// TIA Portal project "FS-DS-09" (V16)
// C100锁螺丝机

(* hardware
DEVICE "S7-1200 station_1"  S7-1200 Station
   slot 0: "Rack_0"  S7-1200 Rack  Rack  V1.0
   slot 1: "FS-DS-09"  CPU 1214C DC/DC/DC  6ES7 214-1AG40-0XB0  V4.4
   slot 2: "DI 16/DQ 16x24VDC_1"  6ES7 223-1BL32-0XB0  V2.0
   slot 3: "DI 8/DQ 8x24VDC_1"  6ES7 223-1BH32-0XB0  V2.0
DEVICE "HMI_1"  KTP700 Basic PN
   slot 0: "HMI_1"  KTP700 Basic PN  6AV2 123-2GB03-0AX0  16.0.0.0
   slot 1: "HMI_RT_1"  KTP700 Basic PN  6AV2 123-2GB03-0AX0  16.0.0.0
   slot 5: "HMI_1.IE_CP_1"  PROFINET Interface  16.0.0.0
      slot 1: "PROFINET Interface_1"  PROFINET Interface
         slot 1: "Port_1"  Port
DEVICE "GSD device_1"  GSD.Device.PN
   slot 0: "机架"  Rack  V1.0
   slot 0: "hj6300"  HJ6300-PN-hj6302-2789  HJ6300-PN  -V1.2
      slot 0: "HJ6300-PN-hj6302-2789"  HJ6300-PN-hj6302-2789
      slot 1: "Interface"  Interface
         slot 1: "Port1"  Port1
         slot 2: "Port2"  Port2
      slot 1: "X逻辑输入 COM1/addr=2/reg=17410_1"  X逻辑输入 COM1/addr=2/reg=17410
         slot 0: "X逻辑输入 COM1/addr=2/reg=17410"  X逻辑输入 COM1/addr=2/reg=17410
      slot 2: "Y逻辑输入 COM1/addr=3/reg=17410_1"  Y逻辑输入 COM1/addr=3/reg=17410
         slot 0: "Y逻辑输入 COM1/addr=3/reg=17410"  Y逻辑输入 COM1/addr=3/reg=17410
      slot 3: "Z逻辑输入 COM1/addr=4/reg=17410_1"  Z逻辑输入 COM1/addr=4/reg=17410
         slot 0: "Z逻辑输入 COM1/addr=4/reg=17410"  Z逻辑输入 COM1/addr=4/reg=17410
      slot 4: "x读取错误编号 COM1/addr=2/reg=24577_1"  x读取错误编号 COM1/addr=2/reg=24577
         slot 0: "x读取错误编号 COM1/addr=2/reg=24577"  x读取错误编号 COM1/addr=2/reg=24577
      slot 5: "y读取错误编号 COM1/addr=3/reg=24577_1"  y读取错误编号 COM1/addr=3/reg=24577
         slot 0: "y读取错误编号 COM1/addr=3/reg=24577"  y读取错误编号 COM1/addr=3/reg=24577
      slot 6: "z读取错误编号 COM1/addr=4/reg=24577_1"  z读取错误编号 COM1/addr=4/reg=24577
         slot 0: "z读取错误编号 COM1/addr=4/reg=24577"  z读取错误编号 COM1/addr=4/reg=24577
      slot 7: "x读取速度 COM1/addr=2/reg=19718_1"  x读取速度 COM1/addr=2/reg=19718
         slot 0: "x读取速度 COM1/addr=2/reg=19718"  x读取速度 COM1/addr=2/reg=19718
      slot 8: "y读取速度 COM1/addr=3/reg=19718_1"  y读取速度 COM1/addr=3/reg=19718
         slot 0: "y读取速度 COM1/addr=3/reg=19718"  y读取速度 COM1/addr=3/reg=19718
      slot 9: "z读取速度 COM1/addr=4/reg=19718_1"  z读取速度 COM1/addr=4/reg=19718
         slot 0: "z读取速度 COM1/addr=4/reg=19718"  z读取速度 COM1/addr=4/reg=19718
      slot 10: "x轴逻辑输出 COM1/addr=2/reg=17481_1"  x轴逻辑输出 COM1/addr=2/reg=17481
         slot 0: "x轴逻辑输出 COM1/addr=2/reg=17481"  x轴逻辑输出 COM1/addr=2/reg=17481
      slot 11: "y轴逻辑输出 COM1/addr=3/reg=17481_1"  y轴逻辑输出 COM1/addr=3/reg=17481
         slot 0: "y轴逻辑输出 COM1/addr=3/reg=17481"  y轴逻辑输出 COM1/addr=3/reg=17481
      slot 12: "z轴逻辑输出 COM1/addr=4/reg=17481_1"  z轴逻辑输出 COM1/addr=4/reg=17481
         slot 0: "z轴逻辑输出 COM1/addr=4/reg=17481"  z轴逻辑输出 COM1/addr=4/reg=17481
      slot 14: "Alarm Data Module_1"  Alarm Data Module
         slot 0: "Alarm Data SubModule"  Alarm Data SubModule
*)

// ===== PLC "FS-DS-09"  CPU 1214C DC/DC/DC =====

VAR_GLOBAL   // PLC tag table "默认变量表"
   "Clock_Byte" AT %MB0 : Byte;
   "Clock_10Hz" AT %M0.0 : Bool;
   "Clock_5Hz" AT %M0.1 : Bool;
   "Clock_2.5Hz" AT %M0.2 : Bool;
   "Clock_2Hz" AT %M0.3 : Bool;
   "Clock_1.25Hz" AT %M0.4 : Bool;
   "Clock_1Hz" AT %M0.5 : Bool;
   "Clock_0.625Hz" AT %M0.6 : Bool;
   "Clock_0.5Hz" AT %M0.7 : Bool;
   "System_Byte" AT %MB1 : Byte;
   "FirstScan" AT %M1.0 : Bool;
   "DiagStatusUpdate" AT %M1.1 : Bool;
   "AlwaysTRUE" AT %M1.2 : Bool;
   "AlwaysFALSE" AT %M1.3 : Bool;
   "Tag_1" AT %M4.0 : Bool;
   "Tag_2" AT %M6.0 : Bool;
   "Tag_3" AT %M5.0 : Bool;
   "Tag_4" AT %M200.0 : Bool;
   "Tag_5" AT %M200.1 : Bool;
   "Tag_6" AT %M30.0 : Bool;
   "Tag_7" AT %M30.1 : Bool;
   "Tag_8" AT %M60.0 : Bool;
   "Tag_9" AT %M20.0 : Bool;
   "Tag_10" AT %M50.0 : Bool;
   "Tag_11" AT %M50.1 : Bool;
   "Tag_12" AT %M50.2 : Bool;
END_VAR

VAR_GLOBAL   // PLC tag table "输入"
   "操作面板急停" AT %I0.0 : Bool;
   "回原位" AT %I0.1 : Bool;
   "启动按钮" AT %I0.2 : Bool;
   "停止按钮" AT %I0.3 : Bool;
   "手动/自动" AT %I0.4 : Bool;
   "按钮盒急停" AT %I0.5 : Bool;
   "左启动" AT %I0.6 : Bool;
   "右启动" AT %I0.7 : Bool;
   "备用" AT %I1.0 : Bool;
   "光幕" AT %I1.1 : Bool;
   "Y1供料器有料" AT %I1.2 : Bool;
   "Y2供料器有料" AT %I1.3 : Bool;
   "1#工装产品信号" AT %I1.4 : Bool;
   "2#工装产品信号" AT %I1.5 : Bool;
   "气夹气缸到位2" AT %I2.0 : Bool;
   "气夹气缸到位1" AT %I2.1 : Bool;
   "工具错误" AT %I2.2 : Bool;
   "工具拧紧OK" AT %I2.3 : Bool;
   "工具拧紧NG" AT %I2.4 : Bool;
   "工具准备好" AT %I2.5 : Bool;
   "工具运行" AT %I2.6 : Bool;
   "气源压力检测" AT %I2.7 : Bool;
   "光栅屏蔽对射开关" AT %I3.0 : Bool;
   "吸附信号" AT %I3.1 : Bool;
   "电批下压气缸下压信号" AT %I3.2 : Bool;
   "安全门" AT %I3.3 : Bool;
   "回原位中" AT %I3.4 : Bool;
   "回原位完成" AT %I3.5 : Bool;
   "X轴故障报警" AT %I3.6 : Bool;
   "Y轴故障报警" AT %I3.7 : Bool;
   "Z轴故障报警" AT %I4.0 : Bool;
   "运动控制卡完成/释放夹紧气缸" AT %I4.1 : Bool;
   "备用_3" AT %I4.2 : Bool;
   "备用_4" AT %I4.3 : Bool;
   "备用_5" AT %I4.4 : Bool;
   "备用_6" AT %I4.5 : Bool;
   "备用_7" AT %I4.6 : Bool;
   "备用_8" AT %I4.7 : Bool;
END_VAR

VAR_GLOBAL   // PLC tag table "输出"
   "三色灯黄色" AT %Q0.0 : Bool;
   "三色灯绿色" AT %Q0.1 : Bool;
   "三色灯红色" AT %Q0.2 : Bool;
   "三色灯蜂鸣器" AT %Q0.3 : Bool;
   "绿色半球指示灯" AT %Q0.4 : Bool;
   "红色半球指示灯" AT %Q0.5 : Bool;
   "运动控制卡任务选择1" AT %Q0.6 : Bool;
   "运动控制卡任务选择2" AT %Q0.7 : Bool;
   "运动控制卡任务选择3" AT %Q1.0 : Bool;
   "运动控制卡任务选择4" AT %Q1.1 : Bool;
   "运动控制卡任务选择5" AT %Q2.0 : Bool;
   "Y1供料器有料输出" AT %Q2.1 : Bool;
   "Y2供料器有料输出" AT %Q2.2 : Bool;
   "运动控制卡启动" AT %Q2.3 : Bool;
   "运动控制卡复位" AT %Q2.4 : Bool;
   "运动控制卡紧急停止" AT %Q2.5 : Bool;
   "运动控制卡停止" AT %Q2.6 : Bool;
   "吸取螺丝电磁阀" AT %Q2.7 : Bool;
   "下压气缸电磁阀" AT %Q3.0 : Bool;
   "工装电磁铁" AT %Q3.1 : Bool;
   "光栅报警" AT %Q3.2 : Bool;
   "伺服复位" AT %Q3.3 : Bool;
   "电批急停" AT %Q3.4 : Bool;
   "电批测试启动" AT %Q3.5 : Bool;
   "FFU" AT %Q3.6 : Bool;
   "照明" AT %Q3.7 : Bool;
   "左启动指示灯" AT %Q4.0 : Bool;
   "右启动指示灯" AT %Q4.1 : Bool;
   "夹紧气缸夹紧" AT %Q4.2 : Bool;
   "伺服报警" AT %Q4.3 : Bool;
   "备用_5(1)" AT %Q4.4 : Bool;
   "备用_6(1)" AT %Q4.5 : Bool;
   "备用_7(1)" AT %Q4.6 : Bool;
   "备用_8(1)" AT %Q4.7 : Bool;
END_VAR

VAR_GLOBAL   // PLC tag table "伺服变量"
   "负方向x" AT %I6.2 : Bool;
   "正方向x" AT %I6.3 : Bool;
   "准备OKx" AT %I42.0 : Bool;
   "故障报警x" AT %I42.1 : Bool;
   "故障代码x" AT %ID17 : DWord;
   "负方向y" AT %I10.2 : Bool;
   "正方向y" AT %I10.3 : Bool;
   "准备OKy" AT %I46.0 : Bool;
   "故障报警y" AT %I46.1 : Bool;
   "故障代码y" AT %ID21 : DWord;
   "负方向z" AT %I14.2 : Bool;
   "正方向z" AT %I14.3 : Bool;
   "准备OKz" AT %I50.0 : Bool;
   "故障报警z" AT %I50.1 : Bool;
   "故障代码z" AT %ID25 : DWord;
END_VAR

TYPE "hengkong"
   STRUCT
      DATA : Struct
         X轴原位 : Bool;
         Y轴原位 : Bool;
         Z轴原位 : Bool;
         Y1供料器有料 : Bool;
         Y2供料器有料 : Bool;
         备用 : Bool;
         任务选择1 : Bool;
         任务选择2 : Bool;
         启动 : Bool;
         回原位 : Bool;
         急停 : Bool;
         OK : Bool;
         光幕和门控报警 : Bool;
         任务选择3 : Bool;
         任务选择4 : Bool;
         任务选择5 : Bool;
         负压传感器 : Bool;
         备用_1 : Bool;
         备用_2 : Bool;
         备用_3 : Bool;
         备用_4 : Bool;
         下压气缸原位 : Bool;
         备用_5 : Bool;
         停止 : Bool;
         吸取螺丝信号 : Bool;
         回原位成功 : Bool;
         回原位中 : Bool;
         下压气缸信号 : Bool;
         备用_6 : Bool;
         认螺帽反转 : Bool;
         备用_7 : Bool;
         备用_8 : Bool;
         任务选择0 : Bool;
         任务选择6 : Bool;
         任务选择7 : Bool;
         备用_9 : Bool;
         启动电批 : Bool;
         备用_10 : Bool;
         备用_11 : Bool;
         备用_12 : Bool;
         获取X轴当前坐标 : LReal;
         获取Y轴当前坐标 : LReal;
         获取Z轴当前坐标 : LReal;
         获取Y2轴当前坐标 : LReal;
         完成螺丝数量 : LReal;
         完成产品数量 : LReal;
         产品合格率 : Word;
         螺丝孔加工完成情况查询 : Word;
         设备报警状态查询 : Word;
         左机加工完成情况查询 : Word;
         右机加工完成情况查询 : Word;
         允许运行指令 : Word;
         从机地址 : Word;
         智能电批任务号 : Word;
         电批加工NG时处理指令 : Word;
      END_STRUCT;
   END_STRUCT;
END_TYPE

TYPE "UDPP"
   STRUCT
      加工文件名称 : String;
      加工文件编号 : Int;
      加工螺丝数量 : Int;
   END_STRUCT;
END_TYPE

TYPE "产品"
   STRUCT
      配方 : Struct
         示教器程序号 : Int;
         产品名称 : String;
      END_STRUCT;
   END_STRUCT;
END_TYPE

DATA_BLOCK "count_DB"   // DB18
{ S7_Optimized_Access := 'TRUE' }
VERSION : 0.1
// stored: InstanceOfName count
"count"
BEGIN
END_DATA_BLOCK

// folder: Alarm

DATA_BLOCK "Alarm FB_DB"   // DB5
{ S7_Optimized_Access := 'TRUE' }
VERSION : 0.1
// stored: InstanceOfName Alarm FB
"Alarm FB"
BEGIN
END_DATA_BLOCK

// folder: Control

DATA_BLOCK "Control_DB"   // DB6
{ S7_Optimized_Access := 'TRUE' }
VERSION : 0.1
// stored: InstanceOfName Control FB
"Control FB"
BEGIN
END_DATA_BLOCK

DATA_BLOCK "Start_DB"   // DB9
{ S7_Optimized_Access := 'TRUE' }
VERSION : 0.1
// stored: InstanceOfName Start
"Start"
BEGIN
END_DATA_BLOCK

DATA_BLOCK "吐钉模式"   // DB20
{ S7_Optimized_Access := 'TRUE' }
VERSION : 0.1
   VAR
      吐钉模式 : Bool;
      下压气缸复位信号 : Bool;
      启动就绪 : Bool;
   END_VAR
BEGIN
END_DATA_BLOCK

// folder: DATA

DATA_BLOCK "IO"   // DB1
{ S7_Optimized_Access := 'FALSE' }
VERSION : 0.1
   VAR
      IN : Array[0..40] of Bool;
      OUT : Array[0..40] of Bool;
   END_VAR
BEGIN
   // IN[0] : 操作面板急停
   // IN[1] : 回原位
   // IN[2] : 启动按钮
   // IN[3] : 停止按钮
   // IN[4] : 手动/自动
   // IN[5] : 按钮盒急停
   // IN[6] : 左启动
   // IN[7] : 右启动
   // IN[8] : 备用
   // IN[9] : 光幕
   // IN[10] : Y1供料器有料
   // IN[11] : Y2供料器有料
   // IN[12] : 1#工装产品信号
   // IN[13] : 2#工装产品信号
   // IN[14] : 气夹气缸到位2
   // IN[15] : 气夹气缸到位1
   // IN[16] : 工具错误
   // IN[17] : 工具拧紧OK
   // IN[18] : 工具拧紧NG
   // IN[19] : 工具准备好
   // IN[20] : 工具运行
   // IN[21] : 气源压力检测
   // IN[22] : 光栅屏蔽对射开关
   // IN[23] : 吸附信号
   // IN[24] : 电批下压气缸下压信号
   // IN[25] : 安全门
   // IN[26] : 回原位中
   // IN[27] : 回原位完成
   // IN[28] : X轴故障报警
   // IN[29] : Y轴故障报警
   // IN[30] : Z轴故障报警
   // IN[31] : 运动控制卡完成/释放夹紧气缸
   // IN[32] : 备用_3
   // IN[33] : 备用_4
   // IN[34] : 备用_5
   // IN[35] : 备用_6
   // IN[36] : 备用_7
   // IN[37] : 备用_8
   // OUT[0] : 三色灯黄色
   // OUT[1] : 三色灯绿色
   // OUT[2] : 三色灯红色
   // OUT[3] : 三色灯蜂鸣器
   // OUT[4] : 绿色半球指示灯
   // OUT[5] : 红色半球指示灯
   // OUT[6] : 运动控制卡任务选择1
   // OUT[7] : 运动控制卡任务选择2
   // OUT[8] : 运动控制卡任务选择3
   // OUT[9] : 运动控制卡任务选择4
   // OUT[10] : 运动控制卡任务选择5
   // OUT[11] : Y1供料器有料输出
   // OUT[12] : Y2供料器有料输出
   // OUT[13] : 运动控制卡启动
   // OUT[14] : 运动控制卡复位
   // OUT[15] : 运动控制卡紧急停止
   // OUT[16] : 运动控制卡停止
   // OUT[17] : 吸取螺丝电磁阀
   // OUT[18] : 下压气缸电磁阀
   // OUT[19] : 工装电磁铁
   // OUT[20] : 光栅报警
   // OUT[21] : 伺服复位
   // OUT[22] : 电批急停
   // OUT[23] : 电批测试启动
   // OUT[24] : FFU
   // OUT[25] : 照明
   // OUT[26] : 左启动指示灯
   // OUT[27] : 右启动指示灯
   // OUT[28] : 夹紧气缸夹紧
   // OUT[29] : 伺服报警
   // OUT[30] : 备用_5(1)
   // OUT[31] : 备用_6(1)
   // OUT[32] : 备用_7(1)
   // OUT[33] : 备用_8(1)
END_DATA_BLOCK

DATA_BLOCK "HengKongMC"   // DB2
{ S7_Optimized_Access := 'FALSE' }
VERSION : 0.1
   VAR
      输入 : Struct   // R/W 01/05/0F
         X轴原位 : Bool;   // 4096
         Y轴原位 : Bool;   // 4097
         Z轴原位 : Bool;   // 4098
         X4备用 : Bool;   // 4099
         Y2供料器有料 : Bool;   // 4100
         电批启动 : Bool;   // 4101
         任务选择1 : Bool;   // 4102
         任务选择2 : Bool;   // 4103
         启动 : Bool;   // 4104
         回原位 : Bool;   // 4105
         急停 : Bool;   // 4106
         OK : Bool;   // 4107
         光幕和门控报警 : Bool;   // 4108
         任务选择3 : Bool;   // 4109
         任务选择4 : Bool;   // 4110
         任务选择5 : Bool;   // 4111
         负压传感器 : Bool;   // 4112
         Y1供料器有料 : Bool;   // 4113
         X19 : Bool;   // 4114
         X20 : Bool;   // 4115
         X21 : Bool;   // 4116
         下压气缸原位 : Bool;   // 4117
         X23 : Bool;   // 4118
         停止 : Bool;   // 4119
      END_STRUCT;
      输出 : Struct   // R/W 01/05/0F
         吸取螺丝信号 : Bool;   // 4176
         回原位成功 : Bool;   // 4177
         回原位中 : Bool;   // 4178
         下压气缸信号 : Bool;   // 4179
         Y5 : Bool;   // 4180
         认螺帽反转 : Bool;   // 4181
         运动控制卡完成信号 : Bool;   // 4182
         Y8 : Bool;   // 4183
         任务选择0 : Bool;   // 4184
         任务选择1 : Bool;   // 4185
         任务选择2 : Bool;   // 4186
         Y12 : Bool;   // 4187
         启动电批 : Bool;   // 4188
         Y14 : Bool;   // 4189
         回原位标志位 : Bool;   // 4190
         Y16 : Bool;   // 4191
      END_STRUCT;
      hengkong : Struct   // 运动控制板卡
         获取X轴当前坐标 : LReal;
         获取Y轴当前坐标 : LReal;
         获取Z轴当前坐标 : LReal;
         获取Y2轴当前坐标 : LReal;
         完成螺丝数量 : Int;
         完成产品数量 : Int;
         产品合格率 : Int;
         螺丝孔加工完成情况查询 : Word;
         设备报警状态查询 : Word;
         左机加工完成情况查询 : Word;
         右机加工完成情况查询 : Word;
         报警异常号 : Int;
         光标处运行标志 : Int;
         当前程序所在行号 : Int;
      END_STRUCT;
   END_VAR
BEGIN
END_DATA_BLOCK

DATA_BLOCK "Alarm"   // DB4
{ S7_Optimized_Access := 'FALSE' }
VERSION : 0.1
   VAR
      运动控制板卡螺丝加工完成情况昂查询 : String;
      运动控制板卡设备报警状态查询 : String;
      运动控制板卡报警 : Bool;
      设备气源压力低报警 : Bool;
      面板急停报警 : Bool;
      操作面板急停报警 : Bool;
      安全门报警 : Bool;
      光幕报警 : Bool;
      回原位超时报警 : Bool;
      Y1供料器超时报警 : Bool;
      Y2供料器超时报警 : Bool;
      工装产品检测1无件报警 : Bool;
      工装产品检测2无件报警 : Bool;
      气缸夹紧1夹紧超时 : Bool;
      气缸夹紧2夹紧超时 : Bool;
      丹尼克尔错误报警 : Bool;
      一级报警 : Bool;
      二级报警 : Bool;
      下压气缸故障 : Bool;
      打螺丝延时过小 : Bool;
      真空检测失败 : Bool;
      吸取螺丝失败 : Bool;
      分料超时 : Bool;
      夹紧气缸故障FB运行前未复位 : Bool;
      下压气缸不在原位 : Bool;
      X轴故障报警 : Bool;
      Y轴故障报警 : Bool;
      Z轴故障报警 : Bool;
   END_VAR
BEGIN
END_DATA_BLOCK

DATA_BLOCK "Blocking function"   // DB7
{ S7_Optimized_Access := 'FALSE' }
VERSION : 0.1
   VAR
      Y1供料器报警屏蔽 : Bool;
      Y2供料器报警屏蔽 : Bool;
      工装产品检测1屏蔽 : Bool;
      工装产品检测2屏蔽 : Bool;
      夹紧气缸1夹紧屏蔽 : Bool;
      夹紧气缸2夹紧屏蔽 : Bool;
      上位机屏蔽 : Bool;
      安全门屏蔽 : Bool;
      光幕屏蔽 : Bool;
   END_VAR
BEGIN
END_DATA_BLOCK

DATA_BLOCK "Control"   // DB8
{ S7_Optimized_Access := 'FALSE' }
VERSION : 0.1
   VAR
      MU : Struct
         上位机吸附电磁阀 : Bool;
         上位机下压气缸电磁阀 : Bool;
         上位机停止 : Bool;
         上位机FFU : Bool;
         上位机照明 : Bool;
         上位机夹紧气缸1夹紧 : Bool;
         上位机夹紧气缸2夹紧 : Bool;
         上位机消音 : Bool;
         上位机错误复位 : Bool;
         上位机加工文件选择 : Int;
         上位机加工文件名称 : String;
         上位机启动信号 : Bool;
         上位机屏蔽信号 : Bool;
         上位机电批启动 : Bool;
         上位机回原位按钮 : Bool;
         上位机行号写入 : Bool;
         上位机行号读取 : Bool;
         上位机工装电磁阀启动 : Bool;
         上位机配方写入 : Bool;
         上位机配方读取 : Bool;
         上位机配方下载到PLC : Bool;
         上位机配方编码 : Int;
         OK : Bool;
         NG : Bool;
         扫码SN : String;
      END_STRUCT;
   END_VAR
BEGIN
END_DATA_BLOCK

DATA_BLOCK "HMI"   // DB10
{ S7_Optimized_Access := 'FALSE' }
VERSION : 0.1
   VAR
      MU : Struct
         HMI吸附电磁阀 : Bool;
         HMI下压气缸电磁阀 : Bool;
         HMI停止 : Bool;
         HMIFFU : Bool;
         HMI照明 : Bool;
         HMI夹紧气缸1夹紧 : Bool;
         HMI夹紧气缸2夹紧 : Bool;
         HMI机消音 : Bool;
         HMI伺服错误复位 : Bool;
         HMI加工文件选择 : Int;
         HMI加工文件名称 : String;
         HMI启动信号 : Bool;
         MHI屏蔽信号 : Bool;
         HMI电批启动 : Bool;
         HMI行号写入 : Bool;
         HMI行号读取 : Bool;
         HMI工装电磁铁启动 : Bool;
         HMI配方下载到PLC : Bool;
         "PLC 配方名称" : String;
         "PLC 程序号" : Int;
         PLC螺丝个数 : Int;
         HMI计数器清零 : Bool;
         HMI合格 : Real;
         "HMI 不合格" : Real;
         HMI合格率 : Real;
         "HMI 产品数" : Real;
         "HMI 运行螺丝个数" : Int;
      END_STRUCT;
      运行状态 : Bool;
      "HMI 运行螺丝个数NG" : Int;
      工件完成信号 : Bool;
   END_VAR
BEGIN
END_DATA_BLOCK

DATA_BLOCK "系统时间"   // DB19
{ S7_Optimized_Access := 'TRUE' }
VERSION : 0.1
   VAR RETAIN
      SET : Bool;
      WRDT : DTL;
      RDDT : DTL;
      RET1 : Word;
      RET2 : Word;
   END_VAR
BEGIN
END_DATA_BLOCK

// folder: Mudbus TCP

DATA_BLOCK "modbus data"   // DB12
{ S7_Optimized_Access := 'FALSE' }
VERSION : 0.1
   VAR
      IPV4 : TCON_IP_v4;
      输入 : Struct
         输入信号1 : Bool;
         输入信号2 : Bool;
         输入信号3 : Bool;
         输入信号4 : Bool;
         输入信号5 : Bool;
         输入信号6 : Bool;
         输入信号7 : Bool;
         输入信号8 : Bool;
         输入信号9 : Bool;
         输入信号10 : Bool;
         输入信号11 : Bool;
         输入信号12 : Bool;
         输入信号13 : Bool;
         输入信号14 : Bool;
         输入信号15 : Bool;
         输入信号16 : Bool;
         输入信号17 : Bool;
         输入信号18 : Bool;
         输入信号19 : Bool;
         输入信号20 : Bool;
         输入信号21 : Bool;
         输入信号22 : Bool;
         输入信号23 : Bool;
         输入信号24 : Bool;
         输入信号25 : Bool;
      END_STRUCT;
      输出 : Struct
         输出信号1 : Bool;
         输出信号2 : Bool;
         输出信号3 : Bool;
         输出信号4 : Bool;
         输出信号5 : Bool;
         输出信号6 : Bool;
         输出信号7 : Bool;
         输出信号8 : Bool;
         输出信号9 : Bool;
         输出信号10 : Bool;
         输出信号11 : Bool;
         输出信号12 : Bool;
         输出信号13 : Bool;
         输出信号14 : Bool;
         输出信号15 : Bool;
         输出信号16 : Bool;
      END_STRUCT;
      Static_1 : Struct
         完成产品数量高位 : Word;
         完成产品数量低位 : Word;
         产品合格率 : Word;
         螺丝加工完成情况查询 : Word;
         设备报警状态查询 : Word;
         左加工完成情况查询 : Word;
         右加工完成情况查询 : Word;
         报警异常行号 : Word;
         Static_1 : Struct
            X轴坐标 : DWord;
            Y轴坐标 : DWord;
            Z轴坐标 : DWord;
            Y1轴坐标 : DWord;
            完成螺丝数量高位 : Word;
            "完成螺丝数量低位‘" : Word;
         END_STRUCT;
      END_STRUCT;
      跳转行号 : Struct
         光标处运行标志 : Word;
         当前程序所在行号 : Word;
      END_STRUCT;
      螺丝重打 : Word := 1;
      回原位标志位写入 : Bool := 0;
   END_VAR
BEGIN
   IPV4.InterfaceId := 64;
   IPV4.ID := 16#01;
   IPV4.ActiveEstablished := 1;
   IPV4.RemoteAddress.ADDR[1] := 192;
   IPV4.RemoteAddress.ADDR[2] := 168;
   IPV4.RemoteAddress.ADDR[3] := 1;
   IPV4.RemoteAddress.ADDR[4] := 152;
   IPV4.RemotePort := 502;
END_DATA_BLOCK

DATA_BLOCK "modbus tcp_DB"   // DB13
{ S7_Optimized_Access := 'TRUE' }
VERSION : 0.1
// stored: InstanceOfName modbus tcp
"modbus tcp"
BEGIN
END_DATA_BLOCK

// folder: System blocks/Program resources

DATA_BLOCK "IEC_Counter_0_DB"   // DB17
{ S7_Optimized_Access := 'TRUE' }
AUTHOR : Simatic
FAMILY : IEC
NAME : CNTR
VERSION : 1.0
// stored: InstanceOfName IEC_COUNTER
"IEC_COUNTER"
BEGIN
END_DATA_BLOCK

// folder: 配方

DATA_BLOCK "UDP"   // DB3
{ S7_Optimized_Access := 'FALSE' }
VERSION : 0.1
   VAR
      Static_1 : Array[0..29] of "UDPP";
   END_VAR
BEGIN
   Static_1[0].加工文件编号 := 0;
   Static_1[1].加工文件编号 := 1;
   Static_1[2].加工文件编号 := 2;
   Static_1[3].加工文件编号 := 3;
   Static_1[4].加工文件编号 := 4;
   Static_1[5].加工文件编号 := 5;
   Static_1[6].加工文件编号 := 6;
   Static_1[7].加工文件编号 := 7;
   Static_1[8].加工文件编号 := 8;
   Static_1[9].加工文件编号 := 9;
   Static_1[10].加工文件编号 := 10;
   Static_1[11].加工文件编号 := 11;
   Static_1[12].加工文件编号 := 12;
   Static_1[13].加工文件编号 := 13;
   Static_1[14].加工文件编号 := 14;
   Static_1[15].加工文件编号 := 15;
   Static_1[16].加工文件编号 := 16;
   Static_1[17].加工文件编号 := 17;
   Static_1[18].加工文件编号 := 18;
   Static_1[19].加工文件编号 := 19;
   Static_1[20].加工文件编号 := 20;
   Static_1[21].加工文件编号 := 21;
   Static_1[22].加工文件编号 := 22;
   Static_1[23].加工文件编号 := 23;
   Static_1[24].加工文件编号 := 24;
   Static_1[25].加工文件编号 := 25;
   Static_1[26].加工文件编号 := 26;
   Static_1[27].加工文件编号 := 27;
   Static_1[28].加工文件编号 := 28;
   Static_1[29].加工文件编号 := 29;
END_DATA_BLOCK

DATA_BLOCK "UDPT"   // DB14
{ S7_Optimized_Access := 'FALSE' }
VERSION : 0.1
BEGIN
END_DATA_BLOCK

DATA_BLOCK "CAOZUO"   // DB15
{ S7_Optimized_Access := 'FALSE' }
VERSION : 0.1
   VAR
      READ : Struct
         REQ : Bool;
         RET_VAL : Word;
         BUSY : Bool;
      END_STRUCT;
      WRITE : Struct
         REQ : Bool;
         RET_VAL : Word;
         BUSY : Bool;
      END_STRUCT;
      Index : Int;
   END_VAR
BEGIN
END_DATA_BLOCK

DATA_BLOCK "配方_DB"   // DB16
{ S7_Optimized_Access := 'TRUE' }
VERSION : 0.1
// stored: InstanceOfName 配方
"配方"
BEGIN
END_DATA_BLOCK

// folder: (top level)

ORGANIZATION_BLOCK "Main"   // OB1, LAD, ProgramCycle
TITLE = "Main Program Sweep (Cycle)"
{ S7_Optimized_Access := 'TRUE' }
VERSION : 0.1
   VAR_INPUT
      Initial_Call : Bool;   // Initial call of this OB
      Remanence : Bool;   // =True, if remanent data are available
   END_VAR
BEGIN

REGION Network 1: Data
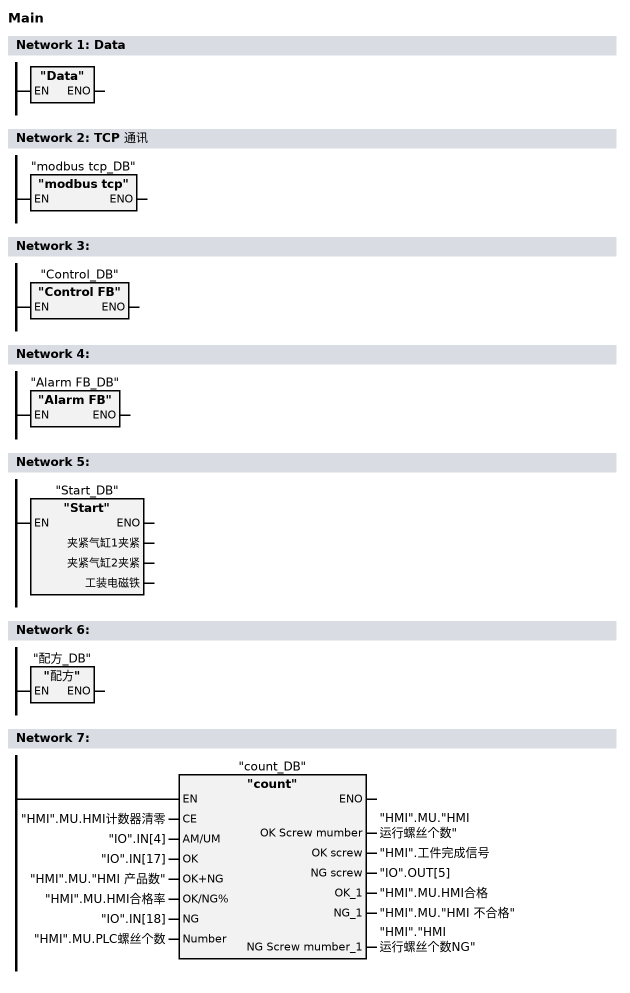
   RUNG wire#powerrail
      "Data"()
   END_RUNG
   // the same network as SCL:
   "Data"();
END_REGION

REGION Network 2: TCP 通讯
   RUNG wire#powerrail
      "modbus tcp_DB"()
   END_RUNG
   // the same network as SCL:
   "modbus tcp_DB"();   // "modbus tcp"
END_REGION

REGION Network 3
   RUNG wire#powerrail
      "Control_DB"()
   END_RUNG
   // the same network as SCL:
   "Control_DB"();   // "Control FB"
END_REGION

REGION Network 4
   RUNG wire#powerrail
      "Alarm FB_DB"()
   END_RUNG
   // the same network as SCL:
   "Alarm FB_DB"();   // "Alarm FB"
END_REGION

REGION Network 5
   RUNG wire#powerrail
      "Start_DB"(夹紧气缸1夹紧 =>, 夹紧气缸2夹紧 =>, 工装电磁铁 =>)
   END_RUNG
   // the same network as SCL:
   "Start_DB"();   // "Start"
END_REGION

REGION Network 6
   RUNG wire#powerrail
      "配方_DB"()
   END_RUNG
   // the same network as SCL:
   "配方_DB"();   // "配方"
END_REGION

REGION Network 7
   RUNG wire#powerrail
      "count_DB"(CE := "HMI".MU.HMI计数器清零, "AM/UM" := "IO".IN[4], OK := "IO".IN[17], "OK+NG" := "HMI".MU."HMI 产品数", "OK/NG%" := "HMI".MU.HMI合格率, NG := "IO".IN[18], Number := "HMI".MU.PLC螺丝个数, "OK Screw mumber" => "HMI".MU."HMI 运行螺丝个数", "OK screw" => "HMI".工件完成信号, "NG screw" => "IO".OUT[5], OK_1 => "HMI".MU.HMI合格, NG_1 => "HMI".MU."HMI 不合格", "NG Screw mumber_1" => "HMI"."HMI 运行螺丝个数NG")
   END_RUNG
   // the same network as SCL:
   "count_DB"(CE := "HMI".MU.HMI计数器清零,   // "count"
              "AM/UM" := "IO".IN[4],
              OK := "IO".IN[17],
              "OK+NG" := "HMI".MU."HMI 产品数",
              "OK/NG%" := "HMI".MU.HMI合格率,
              NG := "IO".IN[18],
              Number := "HMI".MU.PLC螺丝个数,
              "OK Screw mumber" => "HMI".MU."HMI 运行螺丝个数",
              "OK screw" => "HMI".工件完成信号,
              "NG screw" => "IO".OUT[5],
              OK_1 => "HMI".MU.HMI合格,
              NG_1 => "HMI".MU."HMI 不合格",
              "NG Screw mumber_1" => "HMI"."HMI 运行螺丝个数NG");
END_REGION
END_ORGANIZATION_BLOCK

ORGANIZATION_BLOCK "Cyclic interrupt"   // OB30, LAD, CyclicInterrupt
{ S7_Optimized_Access := 'TRUE' }
VERSION : 0.1
   VAR_INPUT
      Initial_Call : Bool;   // Initial call of this OB
      Event_Count : Int;   // Events discarded
   END_VAR
BEGIN

REGION Network 1
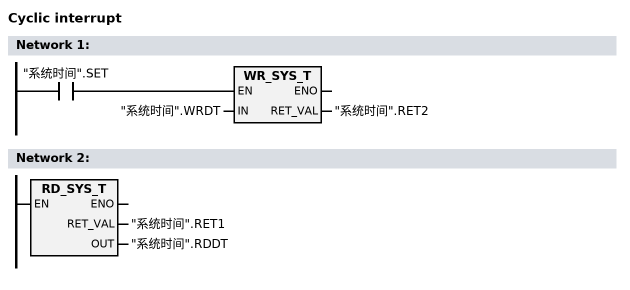
   IF "系统时间".SET THEN "系统时间".RET2 := WR_SYS_T(IN := "系统时间".WRDT); END_IF;
END_REGION

REGION Network 2
   "系统时间".RET1 := RD_SYS_T(OUT => "系统时间".RDDT);
END_REGION
END_ORGANIZATION_BLOCK

// folder: Alarm

FUNCTION_BLOCK "Alarm FB"   // FB3, LAD
{ S7_Optimized_Access := 'TRUE' }
VERSION : 0.1
   VAR
      IEC_Timer_0_Instance : TON_TIME;
      IEC_Timer_0_Instance_1 : TON_TIME;
      IEC_Timer_0_Instance_2 : TON_TIME;
      IEC_Timer_0_Instance_4 : TON_TIME;
      IEC_Timer_0_Instance_3 : TON_TIME;
      报警置位 : Bool;
      蜂鸣器置位 : Bool;
      P1 : Bool;
      R_TRIG_Instance : R_TRIG;
      p2 : Bool;
      p3 : Bool;
      p4 : Bool;
      p5 : Bool;
      p6 : Bool;
      p7 : Bool;
      p8 : Bool;
      p9 : Bool;
      p10 : Bool;
      p11 : Bool;
      p12 : Bool;
      p13 : Bool;
      p14 : Bool;
      p15 : Bool;
   END_VAR
   VAR_TEMP   // added for the SCL form of the ladder/FBD networks
      _w1 : Bool;
      _w2 : Bool;
   END_VAR
BEGIN

REGION Network 1 (SCL): 加工状态情况查询
   IF "HengKongMC".hengkong.螺丝孔加工完成情况查询=0 THEN
       // Statement section IF
       "Alarm".运动控制板卡螺丝加工完成情况昂查询 := '正常';


       ;
   END_IF;//加工状态情况查询
   IF "HengKongMC".hengkong.螺丝孔加工完成情况查询 = 0 THEN
       // Statement section IF
       "Alarm".运动控制板卡螺丝加工完成情况昂查询 := '正常';
       ;
   END_IF;
   IF "HengKongMC".hengkong.螺丝孔加工完成情况查询 = 1 THEN
       // Statement section IF
       "Alarm".运动控制板卡螺丝加工完成情况昂查询 := '拧紧完成';
       ;
   END_IF;
   IF "HengKongMC".hengkong.螺丝孔加工完成情况查询= 16#F4 THEN
       // Statement section IF
       "Alarm".运动控制板卡螺丝加工完成情况昂查询 := '下压气缸故障';
       "Alarm".下压气缸故障 := 1;
   ELSE
       "Alarm".下压气缸故障 := 0;

       ;
   END_IF;
   IF "HengKongMC".hengkong.螺丝孔加工完成情况查询 = 16#F5THEN
       // Statement section IF
       "Alarm".运动控制板卡螺丝加工完成情况昂查询 := '打螺丝完成延时过小';
       "Alarm".打螺丝延时过小 := 1;
   ELSE
       "Alarm".打螺丝延时过小 := 0;
       ;
   END_IF;
   IF "HengKongMC".hengkong.螺丝孔加工完成情况查询 = 16#F6 THEN
       // Statement section IF
       "Alarm".运动控制板卡螺丝加工完成情况昂查询 := '真空检测失败';
       "Alarm".真空检测失败 := 1;
   ELSE
       "Alarm".真空检测失败 := 0;
       ;
   END_IF;
   IF "HengKongMC".hengkong.螺丝孔加工完成情况查询 = 16#F7 THEN
       // Statement section IF
       "Alarm".运动控制板卡螺丝加工完成情况昂查询 := '吸取螺丝失败';
       "Alarm".吸取螺丝失败 := 1;
   ELSE
       "Alarm".吸取螺丝失败 := 0;
       ;
   END_IF;
   IF "HengKongMC".hengkong.螺丝孔加工完成情况查询 = 16#F8 THEN
       // Statement section IF
       "Alarm".运动控制板卡螺丝加工完成情况昂查询 := '分料超时';
       "Alarm".分料超时 := 1;
   ELSE
       "Alarm".分料超时 := 0;

       ;
   END_IF;
   IF"HengKongMC".hengkong.螺丝孔加工完成情况查询 = 16#FA THEN
       // Statement section IF
       "Alarm".运动控制板卡螺丝加工完成情况昂查询 := '夹紧气缸故障FB运行前未复位';
       "Alarm".夹紧气缸故障FB运行前未复位 := 1;
   ELSE
       "Alarm".夹紧气缸故障FB运行前未复位 := 0;

       ;
   END_IF;
   IF "HengKongMC".hengkong.螺丝孔加工完成情况查询 = 16#FC THEN
       // Statement section IF
       "Alarm".运动控制板卡螺丝加工完成情况昂查询 := '下压气缸不在原位';
       "Alarm".下压气缸不在原位 := 1;
   ELSE
       "Alarm".下压气缸不在原位 := 0;
       ;
   END_IF;
   IF "HengKongMC".hengkong.螺丝孔加工完成情况查询 = 16#F8 THEN
       // Statement section IF
       "Alarm".运动控制板卡螺丝加工完成情况昂查询 := '分料超时';
       ;
   END_IF;
   IF "modbus data".Static_1.设备报警状态查询 = 0 THEN
       "Alarm".运动控制板卡设备报警状态查询 := '正常';
   END_IF;
   IF %DB12.DBX29.0  THEN
       // Statement section IF
       "Alarm".运动控制板卡设备报警状态查询 := '急停';
       ;
   END_IF;//设备报警状态查询
   IF  %DB12.DBX29.1  THEN
       // Statement section IF
       "Alarm".运动控制板卡设备报警状态查询  := '光栅';
       ;
   END_IF;
   IF %DB12.DBX29.2  THEN
       // Statement section IF
       "Alarm".运动控制板卡设备报警状态查询  := '伺服报警';
       ;
   END_IF;
   IF %DB12.DBX29.3  THEN
       // Statement section IF
       "Alarm".运动控制板卡设备报警状态查询  := '锁螺丝NG';
       ;
   END_IF;
END_REGION

REGION Network 2 (SCL): 设备报警急停/气源压力低/安全门/工具错误
   "Alarm".操作面板急停报警 := NOT "IO".IN[0];
   "Alarm".设备气源压力低报警 := NOT "IO".IN[21];
   "Alarm".面板急停报警 := NOT "IO".IN[5];
   IF "Blocking function".安全门屏蔽 = 0 THEN
       IF "IO".IN[4] AND "IO".IN[25] = 0 THEN
           "Alarm".安全门报警 := 1;
       ELSE
           "Alarm".安全门报警 := 0;

       END_IF;
       "Alarm".丹尼克尔错误报警 := "IO".IN[16];
   END_IF;

   IF "HengKongMC".hengkong.螺丝孔加工完成情况查询 > 1 OR "HengKongMC".hengkong.设备报警状态查询 > 0 THEN
       // Statement section IF
       "Alarm".运动控制板卡报警 := 1;
   ELSE
       "Alarm".运动控制板卡报警 := 0;
   END_IF;
END_REGION

REGION Network 3 (SCL): 回原位超时报警
   #IEC_Timer_0_Instance(IN:="IO".IN[26],
                         PT:=T#30s,
                         Q=>"Alarm".回原位超时报警);
END_REGION

REGION Network 4: 光幕报警
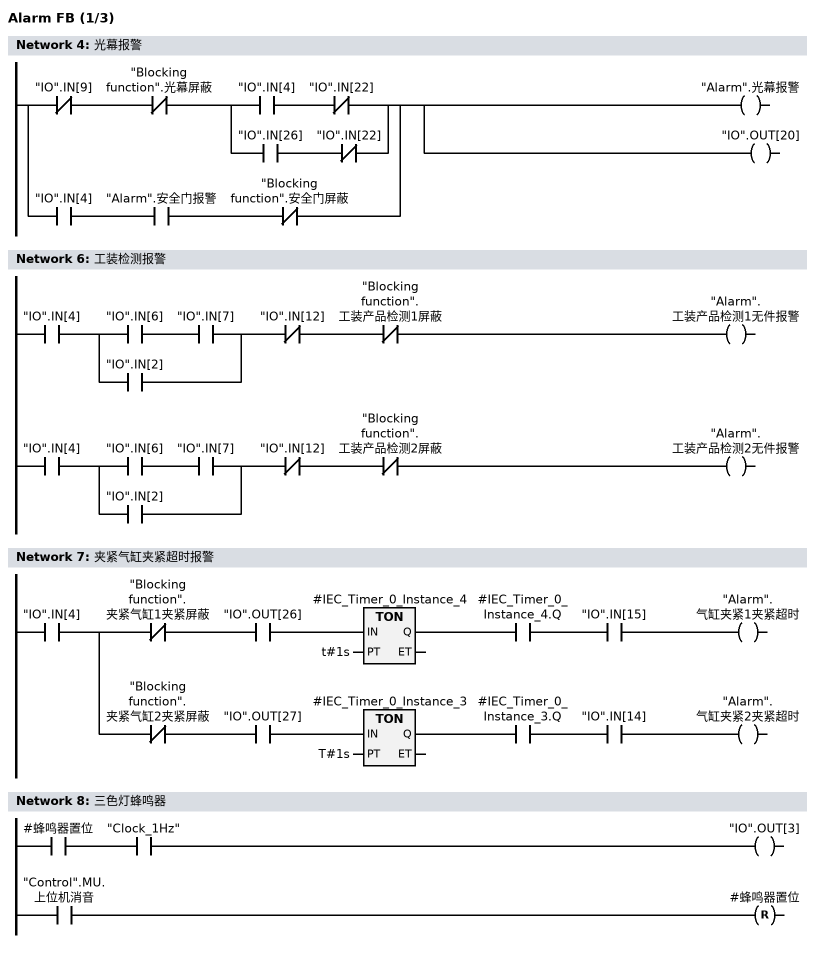
   RUNG wire#powerrail
      I_Contact( "IO".IN[9] )
      I_Contact( "Blocking function".光幕屏蔽 )
      wire#w1
      Contact( "IO".IN[4] )
      I_Contact( "IO".IN[22] )
      wire#w2
      Coil( "Alarm".光幕报警 )
   END_RUNG
   RUNG wire#w1
      Contact( "IO".IN[26] )
      I_Contact( "IO".IN[22] )
   END_RUNG wire#w2
   RUNG wire#powerrail
      Contact( "IO".IN[4] )
      Contact( "Alarm".安全门报警 )
      I_Contact( "Blocking function".安全门屏蔽 )
   END_RUNG wire#w2
   RUNG wire#w2
      Coil( "IO".OUT[20] )
   END_RUNG
   // the same network as SCL:
   "Alarm".光幕报警 := (NOT "IO".IN[9] AND NOT "Blocking function".光幕屏蔽 AND (("IO".IN[4] AND NOT "IO".IN[22]) OR ("IO".IN[26] AND NOT "IO".IN[22]))) OR ("IO".IN[4] AND "Alarm".安全门报警 AND NOT "Blocking function".安全门屏蔽);
   "IO".OUT[20] := "Alarm".光幕报警;
END_REGION

REGION Network 5 (SCL): 供料器超时报警
   IF "Blocking function".Y1供料器报警屏蔽 = 0 THEN
       #IEC_Timer_0_Instance_1(IN := NOT "IO".IN[10],
                               PT := T#5s,
                               Q => "Alarm".Y1供料器超时报警);//Y1 供料器报警
   ELSE
       "Alarm".Y1供料器超时报警 := 0;
   END_IF;//Y1供料器超时报警/屏蔽
   IF "Blocking function".Y2供料器报警屏蔽 = 0 THEN
       #IEC_Timer_0_Instance_2(IN := NOT "IO".IN[11],
                               PT := T#5s,
                               Q => "Alarm".Y2供料器超时报警);//Y2供料器报警
   ELSE
       "Alarm".Y2供料器超时报警 := 0;
   END_IF;//Y2供料器超时报警/屏蔽
END_REGION

REGION Network 6: 工装检测报警
   RUNG wire#powerrail
      Contact( "IO".IN[4] )
      wire#w1
      Contact( "IO".IN[6] )
      Contact( "IO".IN[7] )
      wire#w2
      I_Contact( "IO".IN[12] )
      I_Contact( "Blocking function".工装产品检测1屏蔽 )
      Coil( "Alarm".工装产品检测1无件报警 )
   END_RUNG
   RUNG wire#w1
      Contact( "IO".IN[2] )
   END_RUNG wire#w2
   RUNG wire#powerrail
      Contact( "IO".IN[4] )
      wire#w3
      Contact( "IO".IN[6] )
      Contact( "IO".IN[7] )
      wire#w4
      I_Contact( "IO".IN[12] )
      I_Contact( "Blocking function".工装产品检测2屏蔽 )
      Coil( "Alarm".工装产品检测2无件报警 )
   END_RUNG
   RUNG wire#w3
      Contact( "IO".IN[2] )
   END_RUNG wire#w4
   // the same network as SCL:
   "Alarm".工装产品检测1无件报警 := "IO".IN[4] AND (("IO".IN[6] AND "IO".IN[7]) OR "IO".IN[2]) AND NOT "IO".IN[12] AND NOT "Blocking function".工装产品检测1屏蔽;
   "Alarm".工装产品检测2无件报警 := "IO".IN[4] AND (("IO".IN[6] AND "IO".IN[7]) OR "IO".IN[2]) AND NOT "IO".IN[12] AND NOT "Blocking function".工装产品检测2屏蔽;
END_REGION

REGION Network 7: 夹紧气缸夹紧超时报警
   #IEC_Timer_0_Instance_4(IN := "IO".IN[4] AND NOT "Blocking function".夹紧气缸1夹紧屏蔽 AND "IO".OUT[26], PT := t#1s);   // TON
   "Alarm".气缸夹紧1夹紧超时 := #IEC_Timer_0_Instance_4.Q AND #IEC_Timer_0_Instance_4.Q AND "IO".IN[15];
   #IEC_Timer_0_Instance_3(IN := "IO".IN[4] AND NOT "Blocking function".夹紧气缸2夹紧屏蔽 AND "IO".OUT[27], PT := T#1s);   // TON
   "Alarm".气缸夹紧2夹紧超时 := #IEC_Timer_0_Instance_3.Q AND #IEC_Timer_0_Instance_3.Q AND "IO".IN[14];
END_REGION

REGION Network 8: 三色灯蜂鸣器
   RUNG wire#powerrail
      Contact( #蜂鸣器置位 )
      Contact( "Clock_1Hz" )
      Coil( "IO".OUT[3] )
   END_RUNG
   RUNG wire#powerrail
      Contact( "Control".MU.上位机消音 )
      R_Coil( #蜂鸣器置位 )
   END_RUNG
   // the same network as SCL:
   "IO".OUT[3] := #蜂鸣器置位 AND "Clock_1Hz";
   IF "Control".MU.上位机消音 THEN #蜂鸣器置位 := FALSE; END_IF;
END_REGION

REGION Network 9: 报警
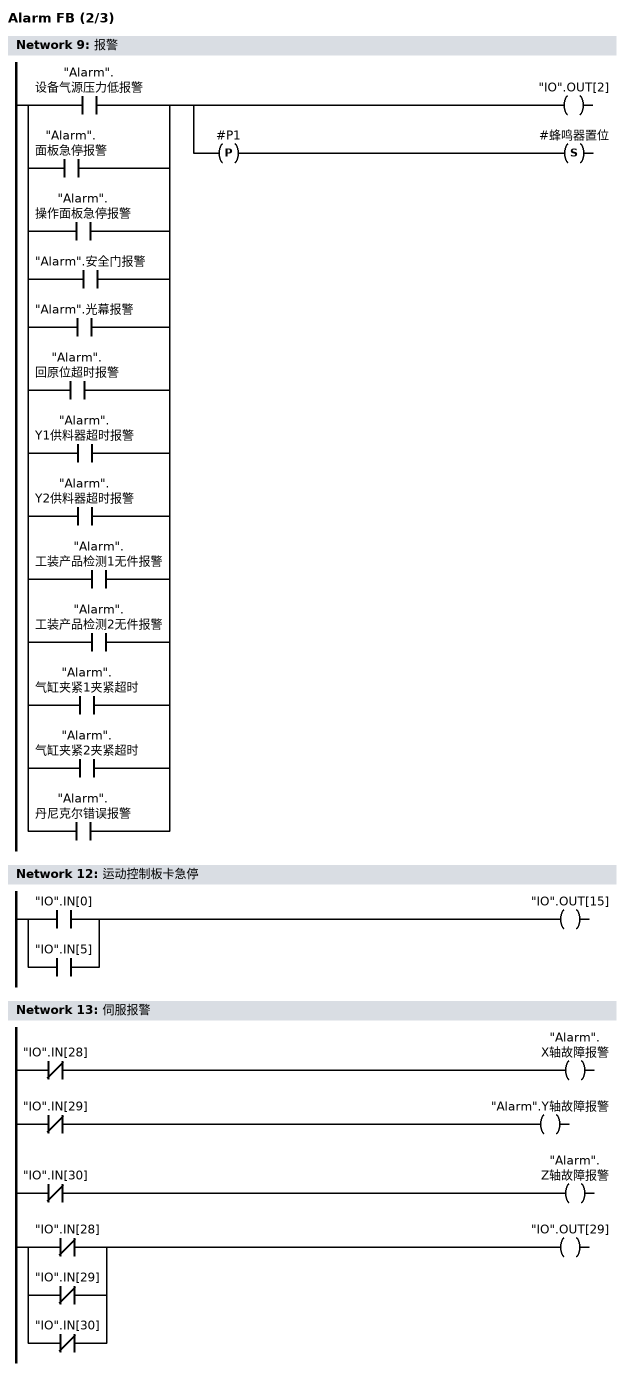
   RUNG wire#powerrail
      Contact( "Alarm".设备气源压力低报警 )
      wire#w1
      Coil( "IO".OUT[2] )
   END_RUNG
   RUNG wire#powerrail
      Contact( "Alarm".面板急停报警 )
   END_RUNG wire#w1
   RUNG wire#powerrail
      Contact( "Alarm".操作面板急停报警 )
   END_RUNG wire#w1
   RUNG wire#powerrail
      Contact( "Alarm".安全门报警 )
   END_RUNG wire#w1
   RUNG wire#powerrail
      Contact( "Alarm".光幕报警 )
   END_RUNG wire#w1
   RUNG wire#powerrail
      Contact( "Alarm".回原位超时报警 )
   END_RUNG wire#w1
   RUNG wire#powerrail
      Contact( "Alarm".Y1供料器超时报警 )
   END_RUNG wire#w1
   RUNG wire#powerrail
      Contact( "Alarm".Y2供料器超时报警 )
   END_RUNG wire#w1
   RUNG wire#powerrail
      Contact( "Alarm".工装产品检测1无件报警 )
   END_RUNG wire#w1
   RUNG wire#powerrail
      Contact( "Alarm".工装产品检测2无件报警 )
   END_RUNG wire#w1
   RUNG wire#powerrail
      Contact( "Alarm".气缸夹紧1夹紧超时 )
   END_RUNG wire#w1
   RUNG wire#powerrail
      Contact( "Alarm".气缸夹紧2夹紧超时 )
   END_RUNG wire#w1
   RUNG wire#powerrail
      Contact( "Alarm".丹尼克尔错误报警 )
   END_RUNG wire#w1
   RUNG wire#w1
      P_Trig( #P1 )
      S_Coil( #蜂鸣器置位 )
   END_RUNG
   // the same network as SCL:
   "IO".OUT[2] := "Alarm".设备气源压力低报警 OR "Alarm".面板急停报警 OR "Alarm".操作面板急停报警 OR "Alarm".安全门报警 OR "Alarm".光幕报警 OR "Alarm".回原位超时报警 OR "Alarm".Y1供料器超时报警 OR "Alarm".Y2供料器超时报警 OR "Alarm".工装产品检测1无件报警 OR "Alarm".工装产品检测2无件报警 OR "Alarm".气缸夹紧1夹紧超时 OR "Alarm".气缸夹紧2夹紧超时 OR "Alarm".丹尼克尔错误报警;
   #_w1 := "Alarm".设备气源压力低报警 OR "Alarm".面板急停报警 OR "Alarm".操作面板急停报警 OR "Alarm".安全门报警 OR "Alarm".光幕报警 OR "Alarm".回原位超时报警 OR "Alarm".Y1供料器超时报警 OR "Alarm".Y2供料器超时报警 OR "Alarm".工装产品检测1无件报警 OR "Alarm".工装产品检测2无件报警 OR "Alarm".气缸夹紧1夹紧超时 OR "Alarm".气缸夹紧2夹紧超时 OR "Alarm".丹尼克尔错误报警;
   #_w2 := #_w1 AND NOT #P1;   // rising edge
   #P1 := #_w1;
   IF #_w2 THEN #蜂鸣器置位 := TRUE; END_IF;
END_REGION

REGION Network 10 (SCL): 一级报警
   IF "Alarm".设备气源压力低报警 OR "Alarm".面板急停报警 OR "Alarm".操作面板急停报警
       OR "Alarm".安全门报警 OR "Alarm".光幕报警 OR "Alarm".回原位超时报警 OR "Alarm".丹尼克尔错误报警 OR "Alarm".X轴故障报警
       OR "Alarm".Y轴故障报警 OR "Alarm".Z轴故障报警
   THEN
       "Alarm".一级报警 := 1;
   ELSE
       "Alarm".一级报警 := 0;
   END_IF;
END_REGION

REGION Network 11 (SCL): 二级报警
   IF "Alarm".回原位超时报警 OR "Alarm".Y1供料器超时报警 OR "Alarm".Y2供料器超时报警 OR "Alarm".工装产品检测1无件报警
       OR "Alarm".工装产品检测2无件报警 OR "Alarm".气缸夹紧1夹紧超时 OR "Alarm".气缸夹紧2夹紧超时 OR "Alarm".下压气缸故障 OR "Alarm".打螺丝延时过小 OR "Alarm".真空检测失败 OR
       "Alarm".吸取螺丝失败 OR "Alarm".分料超时 OR "Alarm".夹紧气缸故障FB运行前未复位 OR "Alarm".下压气缸不在原位 THEN
       "Alarm".二级报警 := 1;
   ELSE
       "Alarm".二级报警 := 0;
   END_IF;
END_REGION

REGION Network 12: 运动控制板卡急停
   RUNG wire#powerrail
      Contact( "IO".IN[0] )
      wire#w1
      Coil( "IO".OUT[15] )
   END_RUNG
   RUNG wire#powerrail
      Contact( "IO".IN[5] )
   END_RUNG wire#w1
   // the same network as SCL:
   "IO".OUT[15] := "IO".IN[0] OR "IO".IN[5];
END_REGION

REGION Network 13: 伺服报警
   RUNG wire#powerrail
      I_Contact( "IO".IN[28] )
      Coil( "Alarm".X轴故障报警 )
   END_RUNG
   RUNG wire#powerrail
      I_Contact( "IO".IN[29] )
      Coil( "Alarm".Y轴故障报警 )
   END_RUNG
   RUNG wire#powerrail
      I_Contact( "IO".IN[30] )
      Coil( "Alarm".Z轴故障报警 )
   END_RUNG
   RUNG wire#powerrail
      I_Contact( "IO".IN[28] )
      wire#w1
      Coil( "IO".OUT[29] )
   END_RUNG
   RUNG wire#powerrail
      I_Contact( "IO".IN[29] )
   END_RUNG wire#w1
   RUNG wire#powerrail
      I_Contact( "IO".IN[30] )
   END_RUNG wire#w1
   // the same network as SCL:
   "Alarm".X轴故障报警 := NOT "IO".IN[28];
   "Alarm".Y轴故障报警 := NOT "IO".IN[29];
   "Alarm".Z轴故障报警 := NOT "IO".IN[30];
   "IO".OUT[29] := NOT "IO".IN[28] OR NOT "IO".IN[29] OR NOT "IO".IN[30];
END_REGION

REGION Network 14: 运动控制板卡急停报警